(* Logix 5000 project; controller FV vendor 1 type 14 code 217 rev 31.11; software revision 31.00; part 58 of 63 *)
(* tags used below, declared in another part *)
   Alarm_Reset : BOOL;
   Always_Off : BOOL;
   Always_On : BOOL;
   CLOCK_system_set : BOOL;
   CLOCKsetvalues : DINT[7];
   CWD : CHECKWORD_FLAGS;
   FV_AV1 : PlantItem;   // AV1
   FV_B100 : INT[255];   // FV FLAGS
   FV_B3 : INT[255];   // BINARY
   FV_B3_0_1_OutputBit : BOOL;
   FV_B50_0_2_StorageBit : BOOL;
   FV_B52 : INT[255];   // WASTE_FLG
   fv_data_file_value_to_move : DINT;
   FV_N12 : INT[255];   // SYS_PARMS System Parameter Fil e
   FV_N50 : INT[255];   // WASTE<PC
   FV_N51 : INT[255];   // WASTE>PC
   FV_N54 : INT[255];   // WASTE_SV
   FV_SFile : INT[255];   // SLC Equivalent System File, So Original Code Can Remain
   FV_T4 : TIMER[10];
   FV_T53 : TIMER[10];
   FV_YSV1_WTX01_AI : PlantItem;   // YSV1_WTX01
   FV_YSV2_WTX01_AI : PlantItem;   // YSV2_WTX01
   FV_YSV2O : PlantItem;   // YSV2O
   FV_YSV3_WTX01_AI : PlantItem;   // YSV3_WTX01
   FV_YSV3O : PlantItem;   // YSV3O
   FV_YSVWaste_AmountAtEnd : REAL;
   One_Minute_One_Scan : BOOL;
   One_Minute_One_Scan_Timer : TIMER;
   One_Second_1_scan : BOOL;
   One_Second_Toggle : BOOL;
   Pitching_transaction_locked_timer : TIMER;
   Pitching_transaction_log : DINT;
   Pitching_transaction_log_delay : DINT;
   Pitching_transaction_log_Done : DINT;
   Pitching_transaction_log_timer : TIMER;
   Reseeding_transaction_locked_timer : TIMER;
   Reseeding_transaction_log : DINT;
   Reseeding_transaction_log_delay : DINT;
   Reseeding_transaction_log_Done : DINT;
   Reseeding_transaction_log_timer : TIMER;
   scada_watchdog : DINT;
   scada_watchdog_tmr : TIMER;
   scada_watchdog_tmr_off : TIMER;
   YSVFilling_transaction_locked_timer : TIMER;
   YSVFilling_transaction_log : DINT;
   YSVFilling_transaction_log_delay : DINT;
   YSVFilling_transaction_log_Done : DINT;
   YSVFilling_transaction_log_timer : TIMER;
(* FV_Common, continued *)

   32: OTL(FV_B52[0].0);
   33: OTL(FV_B52[0].1);
   34: OTL(FV_N51[2].2);
   35: MOV(10,FV_N51[1]);
   36: MOV(10,FV_N51[3]);
   37: MOV(-1,FV_N51[16]);
   38: CLR(FV_N50[0]);
   39: MCR();
   // HANDLE STOP BUTTON
   40: XIC(FV_N50[0].2)XIC(FV_N51[2].2)MCR();
   41: OTU(FV_B52[0].1);
   42: OTU(FV_N51[2].2);
   43: OTL(FV_N51[2].3);
   44: OTL(FV_N51[2].4);
   45: MOV(3,FV_N51[0]);
   46: MOV(0,FV_N51[1]);
   47: CLR(FV_N50[0]);
   48: MCR();
   // HANDLE CONTINUE BUTTON
   49: XIC(FV_N50[0].3)XIC(FV_N51[2].3)MCR();
   50: OTL(FV_B52[0].1);
   51: OTL(FV_N51[2].2);
   52: OTU(FV_N51[2].3);
   // Reset process alarm and parameters
   53: OTU(FV_N51[2].4);
   54: FLL(0,FV_N51[4],4);
   55: MOV(2,FV_N51[0]);
   // Set current Step = Restart Step
   56: MOV(FV_N51[3],FV_N51[1]);
   57: CLR(FV_N50[0]);
   58: MCR();
   // HANDLE ABORT BUTTON
   59: XIC(FV_N50[0].4)XIC(FV_N51[2].4)MCR();
   60: OTU(FV_B52[0].0);
   // Restore YSV operation prior to Waste Transfer
   61: JSR(FV_Set_FV_Datafile_Value,3,FV_N51[13],FV_N51[15],0);
   62: CLR(FV_N51[16]);
   63: CLR(FV_N50[0]);
   64: MCR();
   // Copy step number for PC to display if running
   65: XIC(FV_B52[0].1)MOV(FV_N51[1],FV_N51[9]);
END_ROUTINE

ROUTINE FV_YSVWSTE_MC_25   (* ladder *)
   // Run YSV to Waste  command interpreter
   0: JSR(FV_YSVWSTE_CP_26,0);
   // Run YSV to Waste Process If Active
   1: XIC(FV_B52[0].0)JSR(FV_YSVWSTE_PR_27,0);
   // PostScan YSV to Waste Process If not active
   2: XIO(FV_B52[0].0)OSR(FV_B52[0].2,FV_B50_0_2_StorageBit)XIC(FV_B50_0_2_StorageBit)JSR(FV_YSVWSTE_PR_27,0);
END_ROUTINE

ROUTINE FV_YSVWSTE_PR_27   (* ladder *)
   // YSV TO WASTE- STEP 10 - Initialize
   0: XIC(FV_B52[0].1)EQU(FV_N51[1],10)MCR();
   // Set restart step for this process
   1: MOV(10,FV_N51[3]);
   // Make pointer to selected YSV's data file
   2: ADD(FV_N50[1],140,FV_N51[15]);
   // Make pointer to YSV's Attemporation Data File
   3: ADD(FV_N50[1],135,FV_N51[14]);
   // Save YSV volume at start of transfer
   4: JSR(FV_Get_FV_Datafile_Value,2,FV_N51[15],5)MOV(fv_data_file_value_to_move,FV_N51[17]);
   // Advance to next step
   5: MOV(20,FV_N51[1]);
   6: MCR();
   // Request inlet / outlet valve on correct vessel
   7: [EQU(FV_N50[1],1) MOV(FV_YSV1_WTX01_AI.Scaled,FV_YSVWaste_AmountAtEnd) ,EQU(FV_N50[1],2) MOV(FV_YSV2_WTX01_AI.Scaled,FV_YSVWaste_AmountAtEnd) ,EQU(FV_N50[1],3) MOV(FV_YSV3_WTX01_AI.Scaled,FV_YSVWaste_AmountAtEnd) ];
   // YSV TO WASTE - STEP 20 - Transfer to Waste Yeast
   8: XIC(FV_B52[0].1)EQU(FV_N51[1],20)MCR();
   // Set restart step for this process
   9: MOV(20,FV_N51[3]);
   // Request inlet / outlet valve on correct vessel
   10: [EQU(FV_N50[1],1) OTE(FV_AV1.DriveBits.4) ,EQU(FV_N50[1],2) OTE(FV_YSV2O.DriveBits.4) ,EQU(FV_N50[1],3) OTE(FV_YSV3O.DriveBits.4) ];
   // Allow operator to select process end button
   11: OTE(FV_N51[2].5);
   // Advance to next step when End selected
   12: XIC(FV_N50[0].5)MOV(30,FV_N51[1]);
   13: MCR();
   // YSV TO WASTE - STEP 30 - Save Volume Transfered
   14: XIC(FV_B52[0].1)EQU(FV_N51[1],30)MCR();
   // Delay to allow vessel outlet to close and  weight to steady
   15: TON(FV_T53[2],?,?);
   // Calculate and Save volume pitched
   16: XIC(FV_T53[2].DN)JSR(FV_Get_FV_Datafile_Value,2,FV_N51[15],5)SUB(FV_N51[17],fv_data_file_value_to_move,FV_N54[2]);
   17: XIC(FV_T53[2].DN)MOV(40,FV_N51[1]);
   18: MCR();
   // YSV TO WASTE - STEP 40 - Save Data
   19: XIC(FV_B52[0].1)EQU(FV_N51[1],40)MCR();
   // Set YSV operation to state prior to waste transfer
   20: JSR(FV_Set_FV_Datafile_Value,3,FV_N51[13],FV_N51[15],0);
   // Save YSV number which transfered to PC
   21: MOV(FV_N50[1],FV_N54[1]);
   // Set Save data flag to PC
   22: MOV(1,FV_N54[0]);
   23: CLR(FV_N51[16]);
   24: MCR();
   // CHECK FOR ALARM CONDITIONS
   25: XIC(FV_B52[0].1)MCR();
   26: EQU(FV_N50[1],1)XIC(FV_AV1.CW.[CWD.FAULT])OTU(FV_B52[0].1);
   27: GRT(FV_N51[4],0)OTU(FV_B52[0].1);
   28: XIO(FV_B52[0].1)[MOV(4,FV_N51[0]) ,OTU(FV_N51[2].2) ,OTL(FV_N51[2].3) ,OTL(FV_N51[2].4) ,MOV(0,FV_N51[1]) ];
   29: MCR();
END_ROUTINE

ROUTINE general_timers   (* ladder *)
   0: OTE(Always_On);
   1: XIO(Always_On)OTE(Always_Off);
   2: [XIO(One_Minute_One_Scan_Timer.DN) TON(One_Minute_One_Scan_Timer,?,?) ,XIC(One_Minute_One_Scan_Timer.DN) OTE(One_Minute_One_Scan) ];
   3: XIC(One_Second_1_scan)[ADD(1,scada_watchdog,scada_watchdog) ,GEQ(scada_watchdog,100) CLR(scada_watchdog) ];
   4: [[XIO(One_Second_Toggle) TON(scada_watchdog_tmr,?,?) ,XIC(scada_watchdog_tmr.DN) OTL(One_Second_Toggle) ] ,[XIC(One_Second_Toggle) TON(scada_watchdog_tmr_off,?,?) ,XIC(scada_watchdog_tmr_off.DN) OTU(One_Second_Toggle) ] ];
END_ROUTINE

ROUTINE MainRoutine   (* ladder *)
   0: XIC(s:fs)JSR(Constants,0);
   1: JSR(ClockRoutines,0);
   2: JSR(general_timers,0);
   3: JSR(FV_Analogs,0);
   4: JSR(FV_Move_Temps_To_DataFiles,0);
   // Always Force Alarm Reset to be pushed Until Delphi Code Removed, Original Delphi did not have global alarm reset.
   5: OTU(Alarm_Reset);
   6: JSR(FV_Valves,0);
   7: JSR(FV_Pumps,0);
   8: JSR(FV_Digital_Inputs,0);
   9: JSR(FV_Digital_Outputs,0);
   10: JSR(FV_Old_Checkword_Relaying,0);
   11: JSR(A_FactoryTalk_Requirements,0);
   12: JSR(FV_A_Alarms_From_PLC,0);
   13: JSR(FV_A_Events_From_Scada_IDs,0)JSR(FV_A_Events_From_Scada,0);
   // Fullers FV Control System Fullers FV Aging Control System, ABM Ltd
   // Request Time / Data From Scada on Restart
   14: [XIC(S:FS) ,EQU(FV_SFile[41],0) ]AFI()OTL(FV_N12[0].0);
   15: XIO(FV_N12[0].0)OSR(FV_B3[0].1,FV_B3_0_1_OutputBit)XIC(FV_B3_0_1_OutputBit)[MOV(FV_N12[26],CLOCKsetvalues[0]) MOV(FV_N12[27],CLOCKsetvalues[1]) MOV(FV_N12[28],CLOCKsetvalues[2]) ,MOV(FV_N12[29],CLOCKsetvalues[3]) MOV(FV_N12[30],CLOCKsetvalues[4]) MOV(FV_N12[31],CLOCKsetvalues[5]) ,CLR(CLOCKsetvalues[6]) ,OTL(CLOCK_system_set) ];
   16: XIO(FV_B100[0].3)EQU(FV_SFile[40],FV_N12[35])EQU(FV_SFile[41],FV_N12[36])OTL(FV_B100[0].3);
   // General purpuse 1 second pulse timer
   17: XIC(FV_B100[0].3)EQU(FV_SFile[40],FV_N12[37])EQU(FV_SFile[41],FV_N12[38])OTU(FV_B100[0].3);
   // Communicate I/O with remote devices.
   18: XIO(FV_T4[2].DN)TON(FV_T4[2],?,?);
   // Communicate with other PLCs
   19: JSR(FV_PLC_COMMS_7,0);
   20: JSR(FV_PLC_COMMS_9,0);
   21: JSR(FV_PLC_COMMS_Write_Replacements,0);
   22: JSR(FV_DEBOUNCE_8,0);
   23: JSR(FV_FILLYSV_MC_10,0);
   24: JSR(FV_PITCH_MC_15,0);
   25: JSR(FV_YSVCIP_MC_20,0);
   26: JSR(FV_YSVWSTE_MC_25,0);
   27: JSR(FV_RESEED_MC_30,0);
   28: JSR(FV_LNCIP_MC_35,0);
   29: JSR(FV_YSTFILL_MC_80,0);
   30: JSR(FV_YSTCIP_MC_84,0);
   31: JSR(FV_YSP_COMMS_88,0);
   32: JSR(FV_FV_MCP_100,0);
   33: JSR(FV_GLYCL_PMPS_110,0);
   34: JSR(FV_YSV_ROUSE_112,0);
   35: JSR(FV_YSV_VOLUME_113,0);
   36: ADD(1,FV_SFile[4],FV_SFile[4])GEQ(FV_SFile[4],65000)CLR(FV_SFile[4]);
   37: NEQ(Pitching_transaction_log_delay,0)TON(Pitching_transaction_log_timer,?,?)XIC(Pitching_transaction_log_timer.DN)[CLR(Pitching_transaction_log_delay) ,MOV(1,Pitching_transaction_log) ];
   // When Transaction Has been logged or timed out clear it.
   38: [EQU(Pitching_transaction_log_Done,0) ,NEQ(Pitching_transaction_log,0) TON(Pitching_transaction_locked_timer,?,?) XIC(Pitching_transaction_locked_timer.DN) ][CLR(Pitching_transaction_log) ,MOV(-1,Pitching_transaction_log_Done) ];
   39: NEQ(Reseeding_transaction_log_delay,0)TON(Reseeding_transaction_log_timer,?,?)XIC(Reseeding_transaction_log_timer.DN)[CLR(Reseeding_transaction_log_delay) ,MOV(1,Reseeding_transaction_log) ];
   // When Transaction Has been logged or timed out clear it.
   40: [EQU(Reseeding_transaction_log_Done,0) ,NEQ(Reseeding_transaction_log,0) TON(Reseeding_transaction_locked_timer,?,?) XIC(Reseeding_transaction_locked_timer.DN) ][CLR(Reseeding_transaction_log) ,MOV(-1,Reseeding_transaction_log_Done) ];
   41: NEQ(YSVFilling_transaction_log_delay,0)TON(YSVFilling_transaction_log_timer,?,?)XIC(YSVFilling_transaction_log_timer.DN)[CLR(YSVFilling_transaction_log_delay) ,MOV(1,YSVFilling_transaction_log) ];
   // When Transaction Has been logged or timed out clear it.
   42: [EQU(YSVFilling_transaction_log_Done,0) ,NEQ(YSVFilling_transaction_log,0) TON(YSVFilling_transaction_locked_timer,?,?) XIC(YSVFilling_transaction_locked_timer.DN) ][CLR(YSVFilling_transaction_log) ,MOV(-1,YSVFilling_transaction_log_Done) ];
END_ROUTINE
END_PROGRAM
